REGION Network 11 (STL)
         A     "MC003_EV";
         A(;
         A(;
         L     "CompALTA-MTA".VRealCmp3;
         L     1;
         ==R;
         );
         A(;
         L     "LectAnalógicasMTA".PresionALTA;
         L     "DBParamCmpALTA-MTA".LMedia1;
         >=R;
         );
         O;
         A(;
         L     "CompALTA-MTA".VRealCmp3;
         L     2;
         ==R;
         );
         A(;
         L     "LectAnalógicasMTA".PresionALTA;
         L     "DBParamCmpALTA-MTA".LMedia2;
         >=R;
         );
         O;
         A(;
         L     "CompALTA-MTA".VRealCmp3;
         L     3;
         ==R;
         );
         A(;
         L     "LectAnalógicasMTA".PresionALTA;
         L     "DBParamCmpALTA-MTA".LMedia3;
         >=R;
         );
         O;
         A(;
         L     "CompALTA-MTA".VRealCmp3;
         L     4;
         ==R;
         );
         A(;
         L     "LectAnalógicasMTA".PresionALTA;
         L     "DBParamCmpALTA-MTA".LMedia4;
         >=R;
         );
         O;
         A(;
         L     "CompALTA-MTA".VRealCmp3;
         L     5;
         ==R;
         );
         A(;
         L     "LectAnalógicasMTA".PresionALTA;
         L     "DBParamCmpALTA-MTA".LMedia5;
         >=R;
         );
         O;
         A(;
         L     "CompALTA-MTA".VRealCmp3;
         L     6;
         ==R;
         );
         A(;
         L     "LectAnalógicasMTA".PresionALTA;
         L     "DBParamCmpALTA-MTA".LMedia6;
         >=R;
         );
         );
         L     S5T#30S;
         SF    "Tag_13";
         NOP   0;
         NOP   0;
         NOP   0;
         A     "Tag_13";
         =     #TEMP0;
END_REGION

REGION Network 12: Accionamiento electrovalvula compresor 3 / Carga compresor de alta (válvula 2) BELLIS
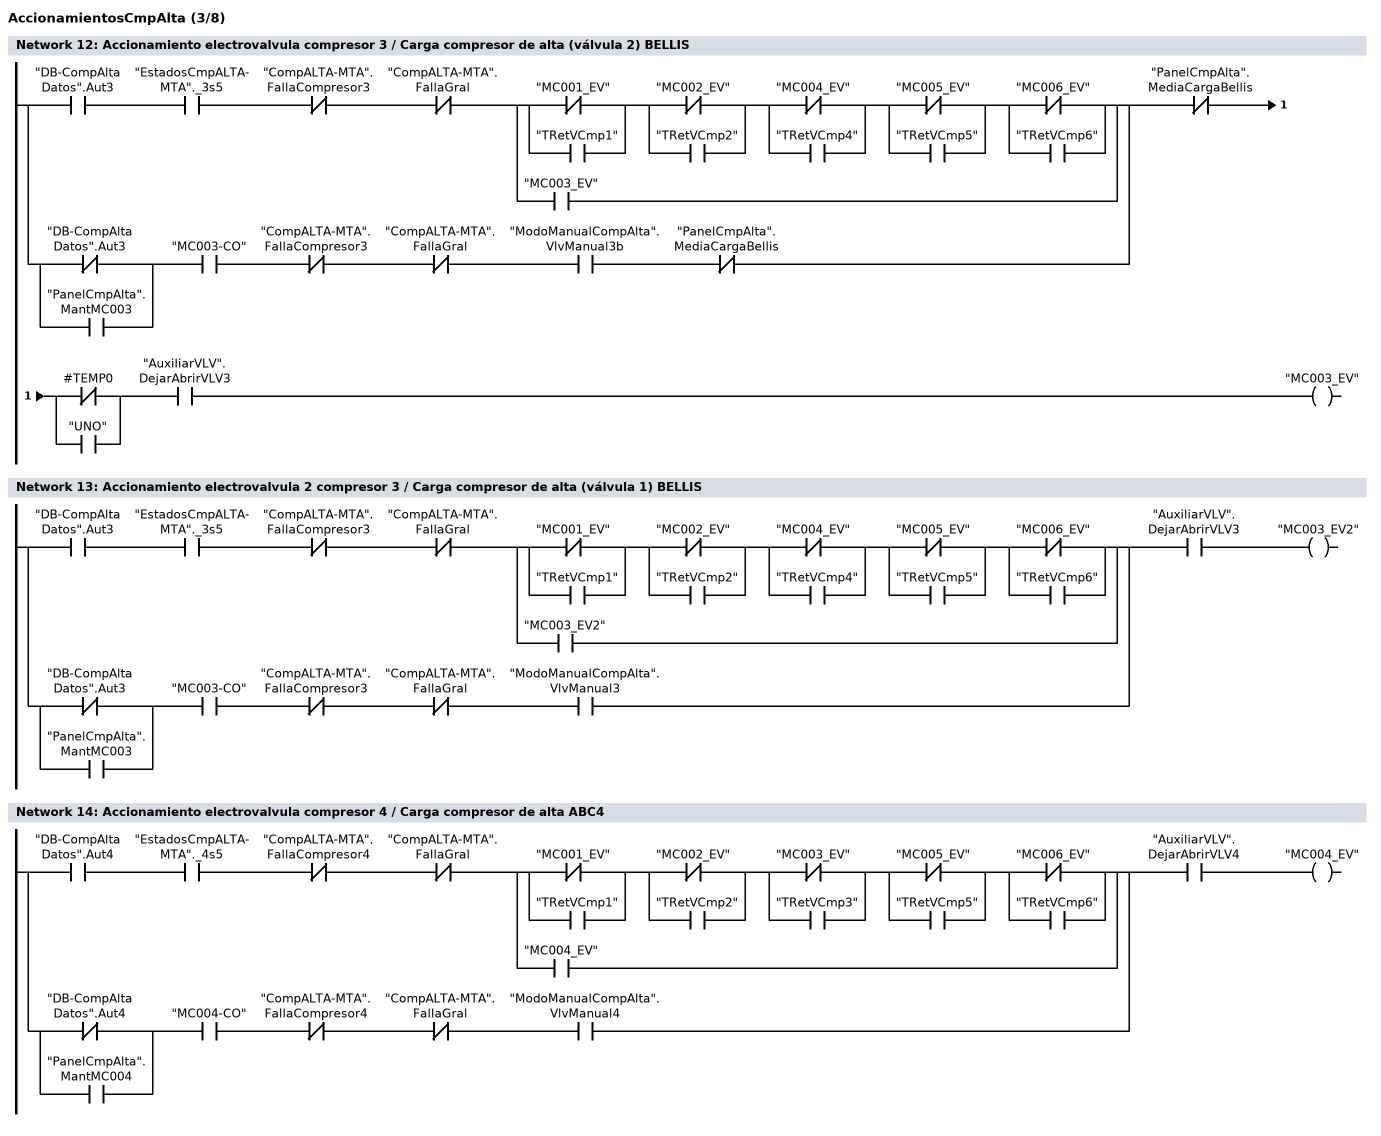
   RUNG wire#powerrail
      Contact( "DB-CompAltaDatos".Aut3 )
      Contact( "EstadosCmpALTA-MTA"._3s5 )
      I_Contact( "CompALTA-MTA".FallaCompresor3 )
      I_Contact( "CompALTA-MTA".FallaGral )
      wire#w1
      I_Contact( "MC001_EV" )
      wire#w2
      I_Contact( "MC002_EV" )
      wire#w3
      I_Contact( "MC004_EV" )
      wire#w4
      I_Contact( "MC005_EV" )
      wire#w5
      I_Contact( "MC006_EV" )
      wire#w6
      I_Contact( "PanelCmpAlta".MediaCargaBellis )
      wire#w8
      I_Contact( #TEMP0 )
      wire#w9
      Contact( "AuxiliarVLV".DejarAbrirVLV3 )
      Coil( "MC003_EV" )
   END_RUNG
   RUNG wire#w1
      Contact( "TRetVCmp1" )
   END_RUNG wire#w2
   RUNG wire#w2
      Contact( "TRetVCmp2" )
   END_RUNG wire#w3
   RUNG wire#w3
      Contact( "TRetVCmp4" )
   END_RUNG wire#w4
   RUNG wire#w4
      Contact( "TRetVCmp5" )
   END_RUNG wire#w5
   RUNG wire#w5
      Contact( "TRetVCmp6" )
   END_RUNG wire#w6
   RUNG wire#w1
      Contact( "MC003_EV" )
   END_RUNG wire#w6
   RUNG wire#powerrail
      I_Contact( "DB-CompAltaDatos".Aut3 )
      wire#w7
      Contact( "MC003-CO" )
      I_Contact( "CompALTA-MTA".FallaCompresor3 )
      I_Contact( "CompALTA-MTA".FallaGral )
      Contact( "ModoManualCompAlta".VlvManual3b )
      I_Contact( "PanelCmpAlta".MediaCargaBellis )
   END_RUNG wire#w6
   RUNG wire#powerrail
      Contact( "PanelCmpAlta".MantMC003 )
   END_RUNG wire#w7
   RUNG wire#w8
      Contact( "UNO" )
   END_RUNG wire#w9
   // the same network as SCL:
   "MC003_EV" := (("DB-CompAltaDatos".Aut3 AND "EstadosCmpALTA-MTA"._3s5 AND NOT "CompALTA-MTA".FallaCompresor3 AND NOT "CompALTA-MTA".FallaGral AND (((NOT "MC001_EV" OR "TRetVCmp1") AND (NOT "MC002_EV" OR "TRetVCmp2") AND (NOT "MC004_EV" OR "TRetVCmp4") AND (NOT "MC005_EV" OR "TRetVCmp5") AND (NOT "MC006_EV" OR "TRetVCmp6")) OR "MC003_EV")) OR ((NOT "DB-CompAltaDatos".Aut3 OR "PanelCmpAlta".MantMC003) AND "MC003-CO" AND NOT "CompALTA-MTA".FallaCompresor3 AND NOT "CompALTA-MTA".FallaGral AND "ModoManualCompAlta".VlvManual3b AND NOT "PanelCmpAlta".MediaCargaBellis)) AND NOT "PanelCmpAlta".MediaCargaBellis AND (NOT #TEMP0 OR "UNO") AND "AuxiliarVLV".DejarAbrirVLV3;
END_REGION

REGION Network 13: Accionamiento electrovalvula 2 compresor 3 / Carga compresor de alta (válvula 1) BELLIS
   RUNG wire#powerrail
      Contact( "DB-CompAltaDatos".Aut3 )
      Contact( "EstadosCmpALTA-MTA"._3s5 )
      I_Contact( "CompALTA-MTA".FallaCompresor3 )
      I_Contact( "CompALTA-MTA".FallaGral )
      wire#w1
      I_Contact( "MC001_EV" )
      wire#w2
      I_Contact( "MC002_EV" )
      wire#w3
      I_Contact( "MC004_EV" )
      wire#w4
      I_Contact( "MC005_EV" )
      wire#w5
      I_Contact( "MC006_EV" )
      wire#w6
      Contact( "AuxiliarVLV".DejarAbrirVLV3 )
      Coil( "MC003_EV2" )
   END_RUNG
   RUNG wire#w1
      Contact( "TRetVCmp1" )
   END_RUNG wire#w2
   RUNG wire#w2
      Contact( "TRetVCmp2" )
   END_RUNG wire#w3
   RUNG wire#w3
      Contact( "TRetVCmp4" )
   END_RUNG wire#w4
   RUNG wire#w4
      Contact( "TRetVCmp5" )
   END_RUNG wire#w5
   RUNG wire#w5
      Contact( "TRetVCmp6" )
   END_RUNG wire#w6
   RUNG wire#w1
      Contact( "MC003_EV2" )
   END_RUNG wire#w6
   RUNG wire#powerrail
      I_Contact( "DB-CompAltaDatos".Aut3 )
      wire#w7
      Contact( "MC003-CO" )
      I_Contact( "CompALTA-MTA".FallaCompresor3 )
      I_Contact( "CompALTA-MTA".FallaGral )
      Contact( "ModoManualCompAlta".VlvManual3 )
   END_RUNG wire#w6
   RUNG wire#powerrail
      Contact( "PanelCmpAlta".MantMC003 )
   END_RUNG wire#w7
   // the same network as SCL:
   "MC003_EV2" := (("DB-CompAltaDatos".Aut3 AND "EstadosCmpALTA-MTA"._3s5 AND NOT "CompALTA-MTA".FallaCompresor3 AND NOT "CompALTA-MTA".FallaGral AND (((NOT "MC001_EV" OR "TRetVCmp1") AND (NOT "MC002_EV" OR "TRetVCmp2") AND (NOT "MC004_EV" OR "TRetVCmp4") AND (NOT "MC005_EV" OR "TRetVCmp5") AND (NOT "MC006_EV" OR "TRetVCmp6")) OR "MC003_EV2")) OR ((NOT "DB-CompAltaDatos".Aut3 OR "PanelCmpAlta".MantMC003) AND "MC003-CO" AND NOT "CompALTA-MTA".FallaCompresor3 AND NOT "CompALTA-MTA".FallaGral AND "ModoManualCompAlta".VlvManual3)) AND "AuxiliarVLV".DejarAbrirVLV3;
END_REGION

REGION Network 14: Accionamiento electrovalvula compresor 4 / Carga compresor de alta ABC4
   RUNG wire#powerrail
      Contact( "DB-CompAltaDatos".Aut4 )
      Contact( "EstadosCmpALTA-MTA"._4s5 )
      I_Contact( "CompALTA-MTA".FallaCompresor4 )
      I_Contact( "CompALTA-MTA".FallaGral )
      wire#w1
      I_Contact( "MC001_EV" )
      wire#w2
      I_Contact( "MC002_EV" )
      wire#w3
      I_Contact( "MC003_EV" )
      wire#w4
      I_Contact( "MC005_EV" )
      wire#w5
      I_Contact( "MC006_EV" )
      wire#w6
      Contact( "AuxiliarVLV".DejarAbrirVLV4 )
      Coil( "MC004_EV" )
   END_RUNG
   RUNG wire#w1
      Contact( "TRetVCmp1" )
   END_RUNG wire#w2
   RUNG wire#w2
      Contact( "TRetVCmp2" )
   END_RUNG wire#w3
   RUNG wire#w3
      Contact( "TRetVCmp3" )
   END_RUNG wire#w4
   RUNG wire#w4
      Contact( "TRetVCmp5" )
   END_RUNG wire#w5
   RUNG wire#w5
      Contact( "TRetVCmp6" )
   END_RUNG wire#w6
   RUNG wire#w1
      Contact( "MC004_EV" )
   END_RUNG wire#w6
   RUNG wire#powerrail
      I_Contact( "DB-CompAltaDatos".Aut4 )
      wire#w7
      Contact( "MC004-CO" )
      I_Contact( "CompALTA-MTA".FallaCompresor4 )
      I_Contact( "CompALTA-MTA".FallaGral )
      Contact( "ModoManualCompAlta".VlvManual4 )
   END_RUNG wire#w6
   RUNG wire#powerrail
      Contact( "PanelCmpAlta".MantMC004 )
   END_RUNG wire#w7
   // the same network as SCL:
   "MC004_EV" := (("DB-CompAltaDatos".Aut4 AND "EstadosCmpALTA-MTA"._4s5 AND NOT "CompALTA-MTA".FallaCompresor4 AND NOT "CompALTA-MTA".FallaGral AND (((NOT "MC001_EV" OR "TRetVCmp1") AND (NOT "MC002_EV" OR "TRetVCmp2") AND (NOT "MC003_EV" OR "TRetVCmp3") AND (NOT "MC005_EV" OR "TRetVCmp5") AND (NOT "MC006_EV" OR "TRetVCmp6")) OR "MC004_EV")) OR ((NOT "DB-CompAltaDatos".Aut4 OR "PanelCmpAlta".MantMC004) AND "MC004-CO" AND NOT "CompALTA-MTA".FallaCompresor4 AND NOT "CompALTA-MTA".FallaGral AND "ModoManualCompAlta".VlvManual4)) AND "AuxiliarVLV".DejarAbrirVLV4;
END_REGION

REGION Network 15: Accionamiento electrovalvula compresor 5 / Carga compresor de alta ABC5
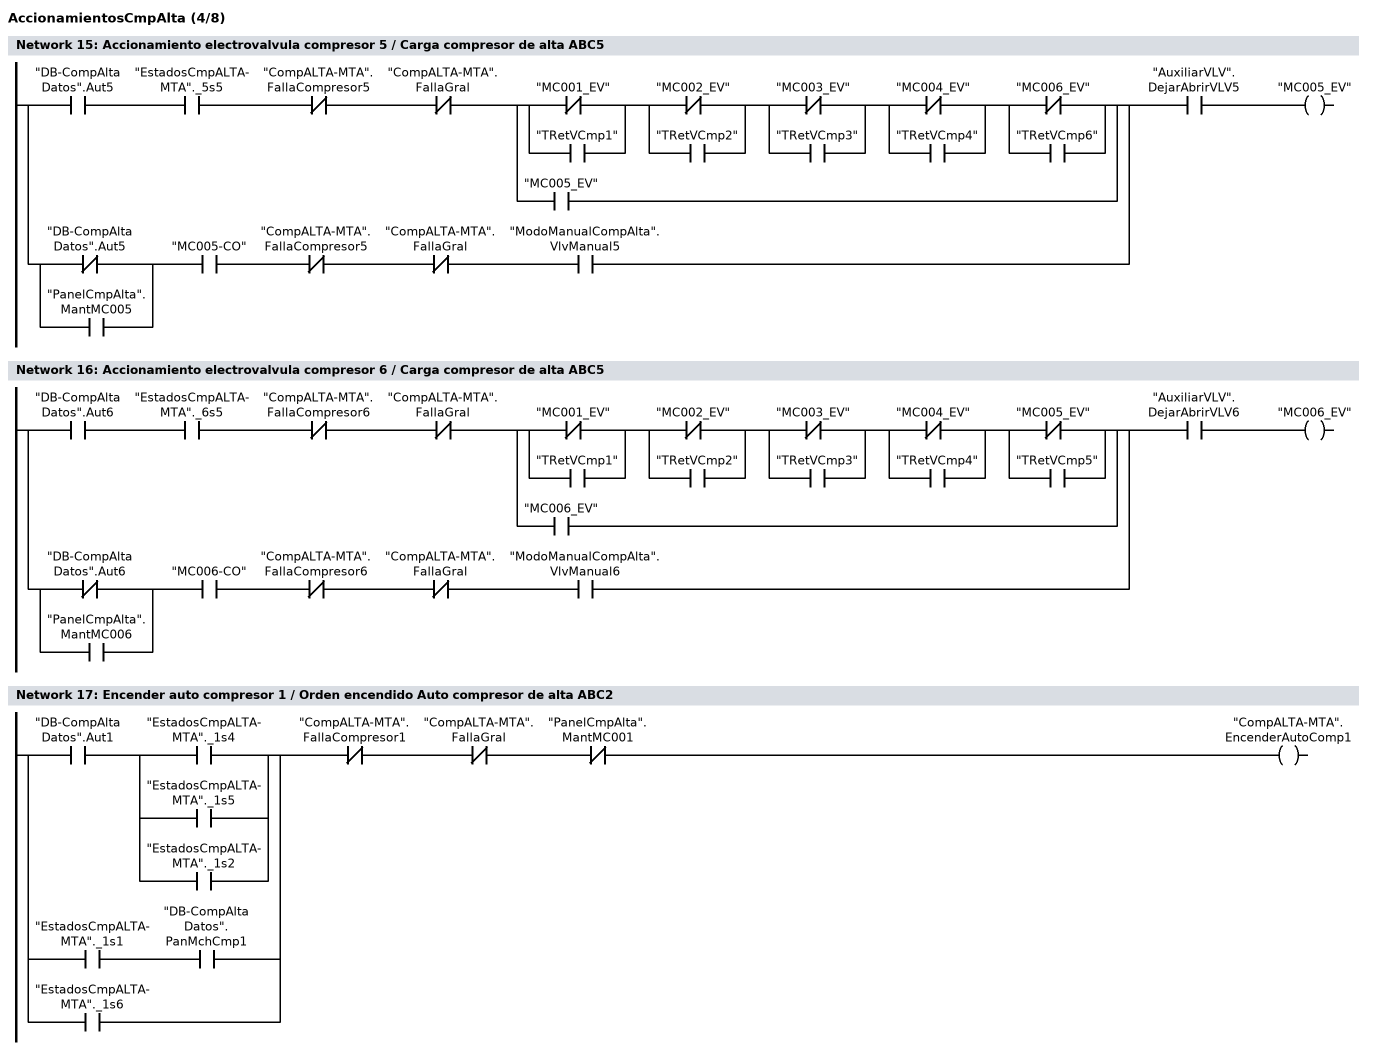
   RUNG wire#powerrail
      Contact( "DB-CompAltaDatos".Aut5 )
      Contact( "EstadosCmpALTA-MTA"._5s5 )
      I_Contact( "CompALTA-MTA".FallaCompresor5 )
      I_Contact( "CompALTA-MTA".FallaGral )
      wire#w1
      I_Contact( "MC001_EV" )
      wire#w2
      I_Contact( "MC002_EV" )
      wire#w3
      I_Contact( "MC003_EV" )
      wire#w4
      I_Contact( "MC004_EV" )
      wire#w5
      I_Contact( "MC006_EV" )
      wire#w6
      Contact( "AuxiliarVLV".DejarAbrirVLV5 )
      Coil( "MC005_EV" )
   END_RUNG
   RUNG wire#w1
      Contact( "TRetVCmp1" )
   END_RUNG wire#w2
   RUNG wire#w2
      Contact( "TRetVCmp2" )
   END_RUNG wire#w3
   RUNG wire#w3
      Contact( "TRetVCmp3" )
   END_RUNG wire#w4
   RUNG wire#w4
      Contact( "TRetVCmp4" )
   END_RUNG wire#w5
   RUNG wire#w5
      Contact( "TRetVCmp6" )
   END_RUNG wire#w6
   RUNG wire#w1
      Contact( "MC005_EV" )
   END_RUNG wire#w6
   RUNG wire#powerrail
      I_Contact( "DB-CompAltaDatos".Aut5 )
      wire#w7
      Contact( "MC005-CO" )
      I_Contact( "CompALTA-MTA".FallaCompresor5 )
      I_Contact( "CompALTA-MTA".FallaGral )
      Contact( "ModoManualCompAlta".VlvManual5 )
   END_RUNG wire#w6
   RUNG wire#powerrail
      Contact( "PanelCmpAlta".MantMC005 )
   END_RUNG wire#w7
   // the same network as SCL:
   "MC005_EV" := (("DB-CompAltaDatos".Aut5 AND "EstadosCmpALTA-MTA"._5s5 AND NOT "CompALTA-MTA".FallaCompresor5 AND NOT "CompALTA-MTA".FallaGral AND (((NOT "MC001_EV" OR "TRetVCmp1") AND (NOT "MC002_EV" OR "TRetVCmp2") AND (NOT "MC003_EV" OR "TRetVCmp3") AND (NOT "MC004_EV" OR "TRetVCmp4") AND (NOT "MC006_EV" OR "TRetVCmp6")) OR "MC005_EV")) OR ((NOT "DB-CompAltaDatos".Aut5 OR "PanelCmpAlta".MantMC005) AND "MC005-CO" AND NOT "CompALTA-MTA".FallaCompresor5 AND NOT "CompALTA-MTA".FallaGral AND "ModoManualCompAlta".VlvManual5)) AND "AuxiliarVLV".DejarAbrirVLV5;
END_REGION

REGION Network 16: Accionamiento electrovalvula compresor 6 / Carga compresor de alta ABC5
   RUNG wire#powerrail
      Contact( "DB-CompAltaDatos".Aut6 )
      Contact( "EstadosCmpALTA-MTA"._6s5 )
      I_Contact( "CompALTA-MTA".FallaCompresor6 )
      I_Contact( "CompALTA-MTA".FallaGral )
      wire#w1
      I_Contact( "MC001_EV" )
      wire#w2
      I_Contact( "MC002_EV" )
      wire#w3
      I_Contact( "MC003_EV" )
      wire#w4
      I_Contact( "MC004_EV" )
      wire#w5
      I_Contact( "MC005_EV" )
      wire#w6
      Contact( "AuxiliarVLV".DejarAbrirVLV6 )
      Coil( "MC006_EV" )
   END_RUNG
   RUNG wire#w1
      Contact( "TRetVCmp1" )
   END_RUNG wire#w2
   RUNG wire#w2
      Contact( "TRetVCmp2" )
   END_RUNG wire#w3
   RUNG wire#w3
      Contact( "TRetVCmp3" )
   END_RUNG wire#w4
   RUNG wire#w4
      Contact( "TRetVCmp4" )
   END_RUNG wire#w5
   RUNG wire#w5
      Contact( "TRetVCmp5" )
   END_RUNG wire#w6
   RUNG wire#w1
      Contact( "MC006_EV" )
   END_RUNG wire#w6
   RUNG wire#powerrail
      I_Contact( "DB-CompAltaDatos".Aut6 )
      wire#w7
      Contact( "MC006-CO" )
      I_Contact( "CompALTA-MTA".FallaCompresor6 )
      I_Contact( "CompALTA-MTA".FallaGral )
      Contact( "ModoManualCompAlta".VlvManual6 )
   END_RUNG wire#w6
   RUNG wire#powerrail
      Contact( "PanelCmpAlta".MantMC006 )
   END_RUNG wire#w7
   // the same network as SCL:
   "MC006_EV" := (("DB-CompAltaDatos".Aut6 AND "EstadosCmpALTA-MTA"._6s5 AND NOT "CompALTA-MTA".FallaCompresor6 AND NOT "CompALTA-MTA".FallaGral AND (((NOT "MC001_EV" OR "TRetVCmp1") AND (NOT "MC002_EV" OR "TRetVCmp2") AND (NOT "MC003_EV" OR "TRetVCmp3") AND (NOT "MC004_EV" OR "TRetVCmp4") AND (NOT "MC005_EV" OR "TRetVCmp5")) OR "MC006_EV")) OR ((NOT "DB-CompAltaDatos".Aut6 OR "PanelCmpAlta".MantMC006) AND "MC006-CO" AND NOT "CompALTA-MTA".FallaCompresor6 AND NOT "CompALTA-MTA".FallaGral AND "ModoManualCompAlta".VlvManual6)) AND "AuxiliarVLV".DejarAbrirVLV6;
END_REGION

REGION Network 17: Encender auto compresor 1 / Orden encendido Auto compresor de alta ABC2
   RUNG wire#powerrail
      Contact( "DB-CompAltaDatos".Aut1 )
      wire#w1
      Contact( "EstadosCmpALTA-MTA"._1s4 )
      wire#w2
      I_Contact( "CompALTA-MTA".FallaCompresor1 )
      I_Contact( "CompALTA-MTA".FallaGral )
      I_Contact( "PanelCmpAlta".MantMC001 )
      Coil( "CompALTA-MTA".EncenderAutoComp1 )
   END_RUNG
   RUNG wire#w1
      Contact( "EstadosCmpALTA-MTA"._1s5 )
   END_RUNG wire#w2
   RUNG wire#w1
      Contact( "EstadosCmpALTA-MTA"._1s2 )
   END_RUNG wire#w2
   RUNG wire#powerrail
      Contact( "EstadosCmpALTA-MTA"._1s1 )
      Contact( "DB-CompAltaDatos".PanMchCmp1 )
   END_RUNG wire#w2
   RUNG wire#powerrail
      Contact( "EstadosCmpALTA-MTA"._1s6 )
   END_RUNG wire#w2
   // the same network as SCL:
   "CompALTA-MTA".EncenderAutoComp1 := (("DB-CompAltaDatos".Aut1 AND ("EstadosCmpALTA-MTA"._1s4 OR "EstadosCmpALTA-MTA"._1s5 OR "EstadosCmpALTA-MTA"._1s2)) OR ("EstadosCmpALTA-MTA"._1s1 AND "DB-CompAltaDatos".PanMchCmp1) OR "EstadosCmpALTA-MTA"._1s6) AND NOT "CompALTA-MTA".FallaCompresor1 AND NOT "CompALTA-MTA".FallaGral AND NOT "PanelCmpAlta".MantMC001;
END_REGION

REGION Network 18: Encender auto compresor 2 / Orden encendido Auto compresor de alta ABC3
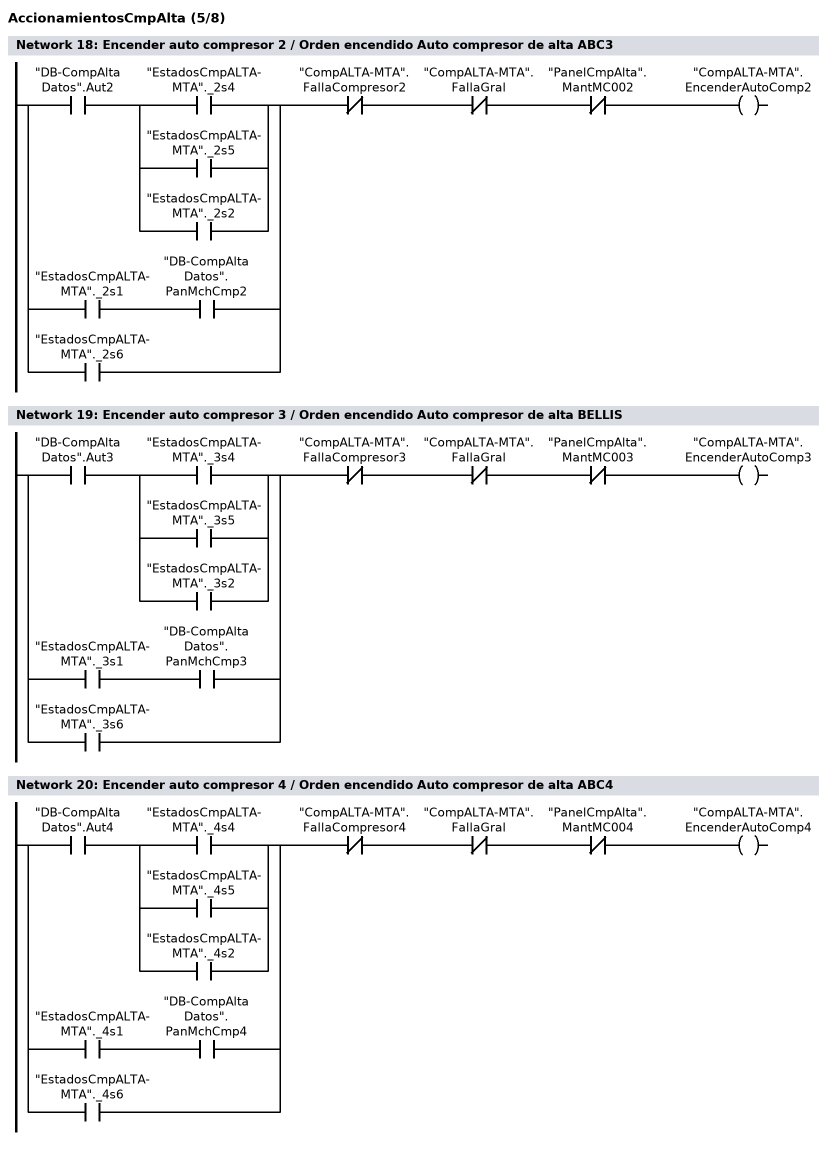
   RUNG wire#powerrail
      Contact( "DB-CompAltaDatos".Aut2 )
      wire#w1
      Contact( "EstadosCmpALTA-MTA"._2s4 )
      wire#w2
      I_Contact( "CompALTA-MTA".FallaCompresor2 )
      I_Contact( "CompALTA-MTA".FallaGral )
      I_Contact( "PanelCmpAlta".MantMC002 )
      Coil( "CompALTA-MTA".EncenderAutoComp2 )
   END_RUNG
   RUNG wire#w1
      Contact( "EstadosCmpALTA-MTA"._2s5 )
   END_RUNG wire#w2
   RUNG wire#w1
      Contact( "EstadosCmpALTA-MTA"._2s2 )
   END_RUNG wire#w2
   RUNG wire#powerrail
      Contact( "EstadosCmpALTA-MTA"._2s1 )
      Contact( "DB-CompAltaDatos".PanMchCmp2 )
   END_RUNG wire#w2
   RUNG wire#powerrail
      Contact( "EstadosCmpALTA-MTA"._2s6 )
   END_RUNG wire#w2
   // the same network as SCL:
   "CompALTA-MTA".EncenderAutoComp2 := (("DB-CompAltaDatos".Aut2 AND ("EstadosCmpALTA-MTA"._2s4 OR "EstadosCmpALTA-MTA"._2s5 OR "EstadosCmpALTA-MTA"._2s2)) OR ("EstadosCmpALTA-MTA"._2s1 AND "DB-CompAltaDatos".PanMchCmp2) OR "EstadosCmpALTA-MTA"._2s6) AND NOT "CompALTA-MTA".FallaCompresor2 AND NOT "CompALTA-MTA".FallaGral AND NOT "PanelCmpAlta".MantMC002;
END_REGION

REGION Network 19: Encender auto compresor 3 / Orden encendido Auto compresor de alta BELLIS
   RUNG wire#powerrail
      Contact( "DB-CompAltaDatos".Aut3 )
      wire#w1
      Contact( "EstadosCmpALTA-MTA"._3s4 )
      wire#w2
      I_Contact( "CompALTA-MTA".FallaCompresor3 )
      I_Contact( "CompALTA-MTA".FallaGral )
      I_Contact( "PanelCmpAlta".MantMC003 )
      Coil( "CompALTA-MTA".EncenderAutoComp3 )
   END_RUNG
   RUNG wire#w1
      Contact( "EstadosCmpALTA-MTA"._3s5 )
   END_RUNG wire#w2
   RUNG wire#w1
      Contact( "EstadosCmpALTA-MTA"._3s2 )
   END_RUNG wire#w2
   RUNG wire#powerrail
      Contact( "EstadosCmpALTA-MTA"._3s1 )
      Contact( "DB-CompAltaDatos".PanMchCmp3 )
   END_RUNG wire#w2
   RUNG wire#powerrail
      Contact( "EstadosCmpALTA-MTA"._3s6 )
   END_RUNG wire#w2
   // the same network as SCL:
   "CompALTA-MTA".EncenderAutoComp3 := (("DB-CompAltaDatos".Aut3 AND ("EstadosCmpALTA-MTA"._3s4 OR "EstadosCmpALTA-MTA"._3s5 OR "EstadosCmpALTA-MTA"._3s2)) OR ("EstadosCmpALTA-MTA"._3s1 AND "DB-CompAltaDatos".PanMchCmp3) OR "EstadosCmpALTA-MTA"._3s6) AND NOT "CompALTA-MTA".FallaCompresor3 AND NOT "CompALTA-MTA".FallaGral AND NOT "PanelCmpAlta".MantMC003;
END_REGION

REGION Network 20: Encender auto compresor 4 / Orden encendido Auto compresor de alta ABC4
   RUNG wire#powerrail
      Contact( "DB-CompAltaDatos".Aut4 )
      wire#w1
      Contact( "EstadosCmpALTA-MTA"._4s4 )
      wire#w2
      I_Contact( "CompALTA-MTA".FallaCompresor4 )
      I_Contact( "CompALTA-MTA".FallaGral )
      I_Contact( "PanelCmpAlta".MantMC004 )
      Coil( "CompALTA-MTA".EncenderAutoComp4 )
   END_RUNG
   RUNG wire#w1
      Contact( "EstadosCmpALTA-MTA"._4s5 )
   END_RUNG wire#w2
   RUNG wire#w1
      Contact( "EstadosCmpALTA-MTA"._4s2 )
   END_RUNG wire#w2
   RUNG wire#powerrail
      Contact( "EstadosCmpALTA-MTA"._4s1 )
      Contact( "DB-CompAltaDatos".PanMchCmp4 )
   END_RUNG wire#w2
   RUNG wire#powerrail
      Contact( "EstadosCmpALTA-MTA"._4s6 )
   END_RUNG wire#w2
   // the same network as SCL:
   "CompALTA-MTA".EncenderAutoComp4 := (("DB-CompAltaDatos".Aut4 AND ("EstadosCmpALTA-MTA"._4s4 OR "EstadosCmpALTA-MTA"._4s5 OR "EstadosCmpALTA-MTA"._4s2)) OR ("EstadosCmpALTA-MTA"._4s1 AND "DB-CompAltaDatos".PanMchCmp4) OR "EstadosCmpALTA-MTA"._4s6) AND NOT "CompALTA-MTA".FallaCompresor4 AND NOT "CompALTA-MTA".FallaGral AND NOT "PanelCmpAlta".MantMC004;
END_REGION

REGION Network 21: Encender auto compresor 5 / Orden encendido Auto compresor de alta ABC5
